// TIA Portal project "EMS" (V15.1) (continued)
   "Carrier_03_SitopSelectStatus" AT %I516.3 : Bool;   // SITOP SELECT STATUS
   "Carrier_03_DCsupplyOnPSCB2" AT %I516.4 : Bool;   // DC SUPPLY ON PSCB 2
   "Carrier_03_SpareInput(4_5)" AT %I516.5 : Bool;   // SPARE INPUT
   "Carrier_03_SpareInput(4_6)" AT %I516.6 : Bool;   // SPARE INPUT
   "Carrier_03_SpareInput(4_7)" AT %I516.7 : Bool;   // SPARE INPUT
   "Carrier_03_PB1_ProdHoldLH" AT %I517.0 : Bool;   // PB 1 PRODUCTION HOLD LH
   "Carrier_03_PB2_ResetLH" AT %I517.1 : Bool;   // PB 2 RESET LH
   "Carrier_03_PB3_ProdHoldRH" AT %I517.2 : Bool;   // PB 3 PRODUCTION HOLD RH
   "Carrier_03_PB4_ResetRH" AT %I517.3 : Bool;   // PB 4 RESET RH
   "Carrier_03_SpareInput(4_14)" AT %I517.4 : Bool;   // SPARE INPUT
   "Carrier_03_SpareInput(4_15)" AT %I517.5 : Bool;   // SPARE INPUT
   "Carrier_03_SpareInput(4_16)" AT %I517.6 : Bool;   // SPARE INPUT
   "Carrier_03_SpareInput(4_17)" AT %I517.7 : Bool;   // SPARE INPUT
   "Carrier_03_Slot5_Output" AT %IW518 : Word;   // SLOT 5 OUTPUT WORD
   "Carrier_03_IRD400_HMI_24VDC_ENABLE" AT %I518.0 : Bool;   // IRD 400 PANEL HMI 24V DC POWER
   "Carrier_03_FaultLight_LH" AT %I518.1 : Bool;   // FAULT LIGHT LH
   "Carrier_03_RunLight_LH" AT %I518.2 : Bool;   // RUN LIGHT LH
   "Carrier_03_FaultLight_RH" AT %I518.3 : Bool;   // FAULT LIGHT RH
   "Carrier_03_RunLight_RH" AT %I518.4 : Bool;   // RUN LIGHT RH
   "Carrier_03_SpareOutput(5_5)" AT %I518.5 : Bool;   // SPARE OUTPUT
   "Carrier_03_SpareOutput(5_6)" AT %I518.6 : Bool;   // SPARE OUTPUT
   "Carrier_03_SpareOutput(5_7)" AT %I518.7 : Bool;   // SPARE OUTPUT
   "Carrier_03_ActualSpeed" AT %IW520 : Word;   // ACTUAL SPEED
   "Carrier_03_CarrierDriveAlarm" AT %IW522 : Word;   // CARRIER DRIVE ALARM
   "Carrier_03_CarrierDriveWarning" AT %IW524 : Word;   // CARRIER DRIVE WARNING
   "Carrier_04_Status" AT %IW550 : Word;   // CARRIER STATUS WORD
   "Carrier_04_Status.0" AT %I550.0 : Bool;   // HEARTBEAT
   "Carrier_04_Status.1" AT %I550.1 : Bool;   // MANUAL
   "Carrier_04_Status.2" AT %I550.2 : Bool;   // IN_AUTO
   "Carrier_04_Status.3" AT %I550.3 : Bool;   // POSITIONING_COMPLETE
   "Carrier_04_Status.4" AT %I550.4 : Bool;   // PRODUCTION HOLD
   "Carrier_04_Status.5" AT %I550.5 : Bool;   // CARRIER MOVING FORWARD
   "Carrier_04_Status.6" AT %I550.6 : Bool;   // CARRIER MOVING REVERSE
   "Carrier_04_Status.7" AT %I550.7 : Bool;   // CARRIER FAULT
   "Carrier_04_Status.8" AT %I551.0 : Bool;   // CRASH DETECT TRIPPED
   "Carrier_04_Status.9" AT %I551.1 : Bool;
   "Carrier_04_Status.10" AT %I551.2 : Bool;
   "Carrier_04_Status.11" AT %I551.3 : Bool;
   "Carrier_04_Status.12" AT %I551.4 : Bool;
   "Carrier_04_Status.13" AT %I551.5 : Bool;
   "Carrier_04_Status.14" AT %I551.6 : Bool;
   "Carrier_04_Status.15" AT %I551.7 : Bool;
   "Carrier_04_SDCFaultCode" AT %IW552 : Word;   // SDC FAULT CODE
   "Carrier_04_CarrierPosition" AT %ID554 : DWord;   // CARRIER POSITION
   "Carrier_04_CarrierNumber" AT %IW558 : Word;   // CARRIER NUMBER
   "Carrier_04_G120DControlWord" AT %IW560 : Word;   // G120D_STW1_CONTROL
   "Carrier_04_G120DControlWord.0" AT %I560.0 : Bool;   // Bit_00_ON
   "Carrier_04_G120DControlWord.1" AT %I560.1 : Bool;   // Bit_01_AUS2_INH
   "Carrier_04_G120DControlWord.2" AT %I560.2 : Bool;   // Bit_02_AUS3_STOP
   "Carrier_04_G120DControlWord.3" AT %I560.3 : Bool;   // Bit_03_EN
   "Carrier_04_G120DControlWord.4" AT %I560.4 : Bool;   // Bit_04_EN_RAMP
   "Carrier_04_G120DControlWord.5" AT %I560.5 : Bool;   // Bit_05_START_RAMP
   "Carrier_04_G120DControlWord.6" AT %I560.6 : Bool;   // Bit_06_SETPOINT
   "Carrier_04_G120DControlWord.7" AT %I560.7 : Bool;   // Bit_07_RESET
   "Carrier_04_G120DControlWord.8" AT %I561.0 : Bool;   // Bit_08_JOG_R
   "Carrier_04_G120DControlWord.9" AT %I561.1 : Bool;   // Bit_09_JOG_L
   "Carrier_04_G120DControlWord.10" AT %I561.2 : Bool;   // Bit_10_CONTR_PLC
   "Carrier_04_G120DControlWord.11" AT %I561.3 : Bool;   // Bit_11_REVERSE
   "Carrier_04_G120DControlWord.12" AT %I561.4 : Bool;   // Bit_12_BRAKE_RELEASE
   "Carrier_04_G120DControlWord.13" AT %I561.5 : Bool;   // Bit_13_DDS
   "Carrier_04_G120DControlWord.14" AT %I561.6 : Bool;   // Bit_14_DO0
   "Carrier_04_G120DControlWord.15" AT %I561.7 : Bool;   // Bit_15_DO1
   "Carrier_04_G120DStatusWord" AT %IW562 : Word;   // G120D_ZSW1_STATUS
   "Carrier_04_G120DStatusWord.0" AT %I562.0 : Bool;   // Bit_00_READY_RUN
   "Carrier_04_G120DStatusWord.1" AT %I562.1 : Bool;   // Bit_01_READY_ON
   "Carrier_04_G120DStatusWord.2" AT %I562.2 : Bool;   // Bit_02_ENABLE
   "Carrier_04_G120DStatusWord.3" AT %I562.3 : Bool;   // Bit_03_FAULT
   "Carrier_04_G120DStatusWord.4" AT %I562.4 : Bool;   // Bit_04_OFF2
   "Carrier_04_G120DStatusWord.5" AT %I562.5 : Bool;   // Bit_05_OFF3
   "Carrier_04_G120DStatusWord.6" AT %I562.6 : Bool;   // Bit_06_LOCK_OUT
   "Carrier_04_G120DStatusWord.7" AT %I562.7 : Bool;   // Bit_07_WARN
   "Carrier_04_G120DStatusWord.8" AT %I563.0 : Bool;   // Bit_08_NO_DEVIATION
   "Carrier_04_G120DStatusWord.9" AT %I563.1 : Bool;   // Bit_09_CONTR_PLC
   "Carrier_04_G120DStatusWord.10" AT %I563.2 : Bool;   // Bit_10_F_MAX
   "Carrier_04_G120DStatusWord.11" AT %I563.3 : Bool;   // Bit_11_LIMIT_REACHED
   "Carrier_04_G120DStatusWord.12" AT %I563.4 : Bool;   // Bit_12_BRAKE_OPEN
   "Carrier_04_G120DStatusWord.13" AT %I563.5 : Bool;   // Bit_13_NO_OVERTEMP
   "Carrier_04_G120DStatusWord.14" AT %I563.6 : Bool;   // Bit_14_CW_CCW
   "Carrier_04_G120DStatusWord.15" AT %I563.7 : Bool;   // Bit_15_OVERL
   "Carrier_04_Slot2_Input" AT %IW564 : Word;   // SLOT 2 INPUT WORD
   "Carrier_04_CrashDetectSW" AT %I564.0 : Bool;   // CRASH DETECT SW
   "Carrier_04_SpareSafetyInput(2_1)" AT %I564.1 : Bool;   // SPARE SAFETY INPUT
   "Carrier_04_SpareSafetyInput(2_2)" AT %I564.2 : Bool;   // SPARE SAFETY INPUT
   "Carrier_04_SpareSafetyInput(2_3)" AT %I564.3 : Bool;   // SPARE SAFETY INPUT
   "Carrier_04_SpareSafetyInput(2_4)" AT %I564.4 : Bool;   // SPARE SAFETY INPUT
   "Carrier_04_SpareSafetyInput(2_5)" AT %I564.5 : Bool;   // SPARE SAFETY INPUT
   "Carrier_04_SpareSafetyInput(2_6)" AT %I564.6 : Bool;   // SPARE SAFETY INPUT
   "Carrier_04_SpareSafetyInput(2_7)" AT %I564.7 : Bool;   // SPARE SAFETY INPUT
   "Carrier_04_Slot3_SafetyOutput" AT %IW565 : Word;   // SLOT 3 SAFETY OUTPUT WORD
   "Carrier_04_Crash_Detect_OK" AT %I565.0 : Bool;   // CARRIER CRASH DETECT
   "Carrier_04_SpareSafetyOutput(3_1)" AT %I565.1 : Bool;   // SPARE SAFETY OUTPUT
   "Carrier_04_SpareSafetyOutput(3_2)" AT %I565.2 : Bool;   // SPARE SAFETY OUTPUT
   "Carrier_04_SpareSafetyOutput(3_3)" AT %I565.3 : Bool;   // SPARE SAFETY OUTPUT
   "Carrier_04_SpareSafetyOutput(3_4)" AT %I565.4 : Bool;   // SPARE SAFETY OUTPUT
   "Carrier_04_SpareSafetyOutput(3_5)" AT %I565.5 : Bool;   // SPARE SAFETY OUTPUT
   "Carrier_04_SpareSafetyOutput(3_6)" AT %I565.6 : Bool;   // SPARE SAFETY OUTPUT
   "Carrier_04_SpareSafetyOutput(3_7)" AT %I565.7 : Bool;   // SPARE SAFETY OUTPUT
   "Carrier_04_Slot4_Input" AT %IW566 : Word;   // SLOT 4 INPUT WORD
   "Carrier_04_480VPowerOn_MDCB1" AT %I566.0 : Bool;   // 480 VAC POWER ON MDCB 1
   "Carrier_04_SpareInput(4_1)" AT %I566.1 : Bool;   // SPARE INPUT
   "Carrier_04_SpareInput(4_2)" AT %I566.2 : Bool;   // SPARE INPUT
   "Carrier_04_SitopSelectStatus" AT %I566.3 : Bool;   // SITOP SELECT STATUS
   "Carrier_04_DCsupplyOnPSCB2" AT %I566.4 : Bool;   // DC SUPPLY ON PSCB 2
   "Carrier_04_SpareInput(4_5)" AT %I566.5 : Bool;   // SPARE INPUT
   "Carrier_04_SpareInput(4_6)" AT %I566.6 : Bool;   // SPARE INPUT
   "Carrier_04_SpareInput(4_7)" AT %I566.7 : Bool;   // SPARE INPUT
   "Carrier_04_PB1_ProdHoldLH" AT %I567.0 : Bool;   // PB 1 PRODUCTION HOLD LH
   "Carrier_04_PB2_ResetLH" AT %I567.1 : Bool;   // PB 2 RESET LH
   "Carrier_04_PB3_ProdHoldRH" AT %I567.2 : Bool;   // PB 3 PRODUCTION HOLD RH
   "Carrier_04_PB4_ResetRH" AT %I567.3 : Bool;   // PB 4 RESET RH
   "Carrier_04_SpareInput(4_14)" AT %I567.4 : Bool;   // SPARE INPUT
   "Carrier_04_SpareInput(4_15)" AT %I567.5 : Bool;   // SPARE INPUT
   "Carrier_04_SpareInput(4_16)" AT %I567.6 : Bool;   // SPARE INPUT
   "Carrier_04_SpareInput(4_17)" AT %I567.7 : Bool;   // SPARE INPUT
   "Carrier_04_Slot5_Output" AT %IW568 : Word;   // SLOT 5 OUTPUT WORD
   "Carrier_04_IRD400_HMI_24VDC_ENABLE" AT %I568.0 : Bool;   // IRD 400 PANEL HMI 24V DC POWER
   "Carrier_04_FaultLight_LH" AT %I568.1 : Bool;   // FAULT LIGHT LH
   "Carrier_04_RunLight_LH" AT %I568.2 : Bool;   // RUN LIGHT LH
   "Carrier_04_FaultLight_RH" AT %I568.3 : Bool;   // FAULT LIGHT RH
   "Carrier_04_RunLight_RH" AT %I568.4 : Bool;   // RUN LIGHT RH
   "Carrier_04_SpareOutput(5_5)" AT %I568.5 : Bool;   // SPARE OUTPUT
   "Carrier_04_SpareOutput(5_6)" AT %I568.6 : Bool;   // SPARE OUTPUT
   "Carrier_04_SpareOutput(5_7)" AT %I568.7 : Bool;   // SPARE OUTPUT
   "Carrier_04_ActualSpeed" AT %IW570 : Word;   // ACTUAL SPEED
   "Carrier_04_CarrierDriveAlarm" AT %IW572 : Word;   // CARRIER DRIVE ALARM
   "Carrier_04_CarrierDriveWarning" AT %IW574 : Word;   // CARRIER DRIVE WARNING
   "Carrier_05_Status" AT %IW600 : Word;   // CARRIER STATUS WORD
   "Carrier_05_Status.0" AT %I600.0 : Bool;   // HEARTBEAT
   "Carrier_05_Status.1" AT %I600.1 : Bool;   // MANUAL
   "Carrier_05_Status.2" AT %I600.2 : Bool;   // IN_AUTO
   "Carrier_05_Status.3" AT %I600.3 : Bool;   // POSITIONING_COMPLETE
   "Carrier_05_Status.4" AT %I600.4 : Bool;   // PRODUCTION HOLD
   "Carrier_05_Status.5" AT %I600.5 : Bool;   // CARRIER MOVING FORWARD
   "Carrier_05_Status.6" AT %I600.6 : Bool;   // CARRIER MOVING REVERSE
   "Carrier_05_Status.7" AT %I600.7 : Bool;   // CARRIER FAULT
   "Carrier_05_Status.8" AT %I601.0 : Bool;   // CRASH DETECT TRIPPED
   "Carrier_05_Status.9" AT %I601.1 : Bool;
   "Carrier_05_Status.10" AT %I601.2 : Bool;
   "Carrier_05_Status.11" AT %I601.3 : Bool;
   "Carrier_05_Status.12" AT %I601.4 : Bool;
   "Carrier_05_Status.13" AT %I601.5 : Bool;
   "Carrier_05_Status.14" AT %I601.6 : Bool;
   "Carrier_05_Status.15" AT %I601.7 : Bool;
   "Carrier_05_SDCFaultCode" AT %IW602 : Word;   // SDC FAULT CODE
   "Carrier_05_CarrierPosition" AT %ID604 : DWord;   // CARRIER POSITION
   "Carrier_05_CarrierNumber" AT %IW608 : Word;   // CARRIER NUMBER
   "Carrier_05_G120DControlWord" AT %IW610 : Word;   // G120D_STW1_CONTROL
   "Carrier_05_G120DControlWord.0" AT %I610.0 : Bool;   // Bit_00_ON
   "Carrier_05_G120DControlWord.1" AT %I610.1 : Bool;   // Bit_01_AUS2_INH
   "Carrier_05_G120DControlWord.2" AT %I610.2 : Bool;   // Bit_02_AUS3_STOP
   "Carrier_05_G120DControlWord.3" AT %I610.3 : Bool;   // Bit_03_EN
   "Carrier_05_G120DControlWord.4" AT %I610.4 : Bool;   // Bit_04_EN_RAMP
   "Carrier_05_G120DControlWord.5" AT %I610.5 : Bool;   // Bit_05_START_RAMP
   "Carrier_05_G120DControlWord.6" AT %I610.6 : Bool;   // Bit_06_SETPOINT
   "Carrier_05_G120DControlWord.7" AT %I610.7 : Bool;   // Bit_07_RESET
   "Carrier_05_G120DControlWord.8" AT %I611.0 : Bool;   // Bit_08_JOG_R
   "Carrier_05_G120DControlWord.9" AT %I611.1 : Bool;   // Bit_09_JOG_L
   "Carrier_05_G120DControlWord.10" AT %I611.2 : Bool;   // Bit_10_CONTR_PLC
   "Carrier_05_G120DControlWord.11" AT %I611.3 : Bool;   // Bit_11_REVERSE
   "Carrier_05_G120DControlWord.12" AT %I611.4 : Bool;   // Bit_12_BRAKE_RELEASE
   "Carrier_05_G120DControlWord.13" AT %I611.5 : Bool;   // Bit_13_DDS
   "Carrier_05_G120DControlWord.14" AT %I611.6 : Bool;   // Bit_14_DO0
   "Carrier_05_G120DControlWord.15" AT %I611.7 : Bool;   // Bit_15_DO1
   "Carrier_05_G120DStatusWord" AT %IW612 : Word;   // G120D_ZSW1_STATUS
   "Carrier_05_G120DStatusWord.0" AT %I612.0 : Bool;   // Bit_00_READY_RUN
   "Carrier_05_G120DStatusWord.1" AT %I612.1 : Bool;   // Bit_01_READY_ON
   "Carrier_05_G120DStatusWord.2" AT %I612.2 : Bool;   // Bit_02_ENABLE
   "Carrier_05_G120DStatusWord.3" AT %I612.3 : Bool;   // Bit_03_FAULT
   "Carrier_05_G120DStatusWord.4" AT %I612.4 : Bool;   // Bit_04_OFF2
   "Carrier_05_G120DStatusWord.5" AT %I612.5 : Bool;   // Bit_05_OFF3
   "Carrier_05_G120DStatusWord.6" AT %I612.6 : Bool;   // Bit_06_LOCK_OUT
   "Carrier_05_G120DStatusWord.7" AT %I612.7 : Bool;   // Bit_07_WARN
   "Carrier_05_G120DStatusWord.8" AT %I613.0 : Bool;   // Bit_08_NO_DEVIATION
   "Carrier_05_G120DStatusWord.9" AT %I613.1 : Bool;   // Bit_09_CONTR_PLC
   "Carrier_05_G120DStatusWord.10" AT %I613.2 : Bool;   // Bit_10_F_MAX
   "Carrier_05_G120DStatusWord.11" AT %I613.3 : Bool;   // Bit_11_LIMIT_REACHED
   "Carrier_05_G120DStatusWord.12" AT %I613.4 : Bool;   // Bit_12_BRAKE_OPEN
   "Carrier_05_G120DStatusWord.13" AT %I613.5 : Bool;   // Bit_13_NO_OVERTEMP
   "Carrier_05_G120DStatusWord.14" AT %I613.6 : Bool;   // Bit_14_CW_CCW
   "Carrier_05_G120DStatusWord.15" AT %I613.7 : Bool;   // Bit_15_OVERL
   "Carrier_05_Slot2_Input" AT %IW614 : Word;   // SLOT 2 INPUT WORD
   "Carrier_05_CrashDetectSW" AT %I614.0 : Bool;   // CRASH DETECT SW
   "Carrier_05_SpareSafetyInput(2_1)" AT %I614.1 : Bool;   // SPARE SAFETY INPUT
   "Carrier_05_SpareSafetyInput(2_2)" AT %I614.2 : Bool;   // SPARE SAFETY INPUT
   "Carrier_05_SpareSafetyInput(2_3)" AT %I614.3 : Bool;   // SPARE SAFETY INPUT
   "Carrier_05_SpareSafetyInput(2_4)" AT %I614.4 : Bool;   // SPARE SAFETY INPUT
   "Carrier_05_SpareSafetyInput(2_5)" AT %I614.5 : Bool;   // SPARE SAFETY INPUT
   "Carrier_05_SpareSafetyInput(2_6)" AT %I614.6 : Bool;   // SPARE SAFETY INPUT
   "Carrier_05_SpareSafetyInput(2_7)" AT %I614.7 : Bool;   // SPARE SAFETY INPUT
   "Carrier_05_Slot3_SafetyOutput" AT %IW615 : Word;   // SLOT 3 SAFETY OUTPUT WORD
   "Carrier_05_Crash_Detect_OK" AT %I615.0 : Bool;   // CARRIER CRASH DETECT
   "Carrier_05_SpareSafetyOutput(3_1)" AT %I615.1 : Bool;   // SPARE SAFETY OUTPUT
   "Carrier_05_SpareSafetyOutput(3_2)" AT %I615.2 : Bool;   // SPARE SAFETY OUTPUT
   "Carrier_05_SpareSafetyOutput(3_3)" AT %I615.3 : Bool;   // SPARE SAFETY OUTPUT
   "Carrier_05_SpareSafetyOutput(3_4)" AT %I615.4 : Bool;   // SPARE SAFETY OUTPUT
   "Carrier_05_SpareSafetyOutput(3_5)" AT %I615.5 : Bool;   // SPARE SAFETY OUTPUT
   "Carrier_05_SpareSafetyOutput(3_6)" AT %I615.6 : Bool;   // SPARE SAFETY OUTPUT
   "Carrier_05_SpareSafetyOutput(3_7)" AT %I615.7 : Bool;   // SPARE SAFETY OUTPUT
   "Carrier_05_Slot4_Input" AT %IW616 : Word;   // SLOT 4 INPUT WORD
   "Carrier_05_480VPowerOn_MDCB1" AT %I616.0 : Bool;   // 480 VAC POWER ON MDCB 1
   "Carrier_05_SpareInput(4_1)" AT %I616.1 : Bool;   // SPARE INPUT
   "Carrier_05_SpareInput(4_2)" AT %I616.2 : Bool;   // SPARE INPUT
   "Carrier_05_SitopSelectStatus" AT %I616.3 : Bool;   // SITOP SELECT STATUS
   "Carrier_05_DCsupplyOnPSCB2" AT %I616.4 : Bool;   // DC SUPPLY ON PSCB 2
   "Carrier_05_SpareInput(4_5)" AT %I616.5 : Bool;   // SPARE INPUT
   "Carrier_05_SpareInput(4_6)" AT %I616.6 : Bool;   // SPARE INPUT
   "Carrier_05_SpareInput(4_7)" AT %I616.7 : Bool;   // SPARE INPUT
   "Carrier_05_PB1_ProdHoldLH" AT %I617.0 : Bool;   // PB 1 PRODUCTION HOLD LH
   "Carrier_05_PB2_ResetLH" AT %I617.1 : Bool;   // PB 2 RESET LH
   "Carrier_05_PB3_ProdHoldRH" AT %I617.2 : Bool;   // PB 3 PRODUCTION HOLD RH
   "Carrier_05_PB4_ResetRH" AT %I617.3 : Bool;   // PB 4 RESET RH
   "Carrier_05_SpareInput(4_14)" AT %I617.4 : Bool;   // SPARE INPUT
   "Carrier_05_SpareInput(4_15)" AT %I617.5 : Bool;   // SPARE INPUT
   "Carrier_05_SpareInput(4_16)" AT %I617.6 : Bool;   // SPARE INPUT
   "Carrier_05_SpareInput(4_17)" AT %I617.7 : Bool;   // SPARE INPUT
   "Carrier_05_Slot5_Output" AT %IW618 : Word;   // SLOT 5 OUTPUT WORD
   "Carrier_05_IRD400_HMI_24VDC_ENABLE" AT %I618.0 : Bool;   // IRD 400 PANEL HMI 24V DC POWER
   "Carrier_05_FaultLight_LH" AT %I618.1 : Bool;   // FAULT LIGHT LH
   "Carrier_05_RunLight_LH" AT %I618.2 : Bool;   // RUN LIGHT LH
   "Carrier_05_FaultLight_RH" AT %I618.3 : Bool;   // FAULT LIGHT RH
   "Carrier_05_RunLight_RH" AT %I618.4 : Bool;   // RUN LIGHT RH
   "Carrier_05_SpareOutput(5_5)" AT %I618.5 : Bool;   // SPARE OUTPUT
   "Carrier_05_SpareOutput(5_6)" AT %I618.6 : Bool;   // SPARE OUTPUT
   "Carrier_05_SpareOutput(5_7)" AT %I618.7 : Bool;   // SPARE OUTPUT
   "Carrier_05_ActualSpeed" AT %IW620 : Word;   // ACTUAL SPEED
   "Carrier_05_CarrierDriveAlarm" AT %IW622 : Word;   // CARRIER DRIVE ALARM
   "Carrier_05_CarrierDriveWarning" AT %IW624 : Word;   // CARRIER DRIVE WARNING
   "Carrier_06_Status" AT %IW650 : Word;   // CARRIER STATUS WORD
   "Carrier_06_Status.0" AT %I650.0 : Bool;   // HEARTBEAT
   "Carrier_06_Status.1" AT %I650.1 : Bool;   // MANUAL
   "Carrier_06_Status.2" AT %I650.2 : Bool;   // IN_AUTO
   "Carrier_06_Status.3" AT %I650.3 : Bool;   // POSITIONING_COMPLETE
   "Carrier_06_Status.4" AT %I650.4 : Bool;   // PRODUCTION HOLD
   "Carrier_06_Status.5" AT %I650.5 : Bool;   // CARRIER MOVING FORWARD
   "Carrier_06_Status.6" AT %I650.6 : Bool;   // CARRIER MOVING REVERSE
   "Carrier_06_Status.7" AT %I650.7 : Bool;   // CARRIER FAULT
   "Carrier_06_Status.8" AT %I651.0 : Bool;   // CRASH DETECT TRIPPED
   "Carrier_06_Status.9" AT %I651.1 : Bool;
   "Carrier_06_Status.10" AT %I651.2 : Bool;
   "Carrier_06_Status.11" AT %I651.3 : Bool;
   "Carrier_06_Status.12" AT %I651.4 : Bool;
   "Carrier_06_Status.13" AT %I651.5 : Bool;
   "Carrier_06_Status.14" AT %I651.6 : Bool;
   "Carrier_06_Status.15" AT %I651.7 : Bool;
   "Carrier_06_SDCFaultCode" AT %IW652 : Word;   // SDC FAULT CODE
   "Carrier_06_CarrierPosition" AT %ID654 : DWord;   // CARRIER POSITION
   "Carrier_06_CarrierNumber" AT %IW658 : Word;   // CARRIER NUMBER
   "Carrier_06_G120DControlWord" AT %IW660 : Word;   // G120D_STW1_CONTROL
   "Carrier_06_G120DControlWord.0" AT %I660.0 : Bool;   // Bit_00_ON
   "Carrier_06_G120DControlWord.1" AT %I660.1 : Bool;   // Bit_01_AUS2_INH
   "Carrier_06_G120DControlWord.2" AT %I660.2 : Bool;   // Bit_02_AUS3_STOP
   "Carrier_06_G120DControlWord.3" AT %I660.3 : Bool;   // Bit_03_EN
   "Carrier_06_G120DControlWord.4" AT %I660.4 : Bool;   // Bit_04_EN_RAMP
   "Carrier_06_G120DControlWord.5" AT %I660.5 : Bool;   // Bit_05_START_RAMP
   "Carrier_06_G120DControlWord.6" AT %I660.6 : Bool;   // Bit_06_SETPOINT
   "Carrier_06_G120DControlWord.7" AT %I660.7 : Bool;   // Bit_07_RESET
   "Carrier_06_G120DControlWord.8" AT %I661.0 : Bool;   // Bit_08_JOG_R
   "Carrier_06_G120DControlWord.9" AT %I661.1 : Bool;   // Bit_09_JOG_L
   "Carrier_06_G120DControlWord.10" AT %I661.2 : Bool;   // Bit_10_CONTR_PLC
   "Carrier_06_G120DControlWord.11" AT %I661.3 : Bool;   // Bit_11_REVERSE
   "Carrier_06_G120DControlWord.12" AT %I661.4 : Bool;   // Bit_12_BRAKE_RELEASE
   "Carrier_06_G120DControlWord.13" AT %I661.5 : Bool;   // Bit_13_DDS
   "Carrier_06_G120DControlWord.14" AT %I661.6 : Bool;   // Bit_14_DO0
   "Carrier_06_G120DControlWord.15" AT %I661.7 : Bool;   // Bit_15_DO1
   "Carrier_06_G120DStatusWord" AT %IW662 : Word;   // G120D_ZSW1_STATUS
   "Carrier_06_G120DStatusWord.0" AT %I662.0 : Bool;   // Bit_00_READY_RUN
   "Carrier_06_G120DStatusWord.1" AT %I662.1 : Bool;   // Bit_01_READY_ON
   "Carrier_06_G120DStatusWord.2" AT %I662.2 : Bool;   // Bit_02_ENABLE
   "Carrier_06_G120DStatusWord.3" AT %I662.3 : Bool;   // Bit_03_FAULT
   "Carrier_06_G120DStatusWord.4" AT %I662.4 : Bool;   // Bit_04_OFF2
   "Carrier_06_G120DStatusWord.5" AT %I662.5 : Bool;   // Bit_05_OFF3
   "Carrier_06_G120DStatusWord.6" AT %I662.6 : Bool;   // Bit_06_LOCK_OUT
   "Carrier_06_G120DStatusWord.7" AT %I662.7 : Bool;   // Bit_07_WARN
   "Carrier_06_G120DStatusWord.8" AT %I663.0 : Bool;   // Bit_08_NO_DEVIATION
   "Carrier_06_G120DStatusWord.9" AT %I663.1 : Bool;   // Bit_09_CONTR_PLC
   "Carrier_06_G120DStatusWord.10" AT %I663.2 : Bool;   // Bit_10_F_MAX
   "Carrier_06_G120DStatusWord.11" AT %I663.3 : Bool;   // Bit_11_LIMIT_REACHED
   "Carrier_06_G120DStatusWord.12" AT %I663.4 : Bool;   // Bit_12_BRAKE_OPEN
   "Carrier_06_G120DStatusWord.13" AT %I663.5 : Bool;   // Bit_13_NO_OVERTEMP
   "Carrier_06_G120DStatusWord.14" AT %I663.6 : Bool;   // Bit_14_CW_CCW
   "Carrier_06_G120DStatusWord.15" AT %I663.7 : Bool;   // Bit_15_OVERL
   "Carrier_06_Slot2_Input" AT %IW664 : Word;   // SLOT 2 INPUT WORD
   "Carrier_06_CrashDetectSW" AT %I664.0 : Bool;   // CRASH DETECT SW
   "Carrier_06_SpareSafetyInput(2_1)" AT %I664.1 : Bool;   // SPARE SAFETY INPUT
   "Carrier_06_SpareSafetyInput(2_2)" AT %I664.2 : Bool;   // SPARE SAFETY INPUT
   "Carrier_06_SpareSafetyInput(2_3)" AT %I664.3 : Bool;   // SPARE SAFETY INPUT
   "Carrier_06_SpareSafetyInput(2_4)" AT %I664.4 : Bool;   // SPARE SAFETY INPUT
   "Carrier_06_SpareSafetyInput(2_5)" AT %I664.5 : Bool;   // SPARE SAFETY INPUT
   "Carrier_06_SpareSafetyInput(2_6)" AT %I664.6 : Bool;   // SPARE SAFETY INPUT
   "Carrier_06_SpareSafetyInput(2_7)" AT %I664.7 : Bool;   // SPARE SAFETY INPUT
   "Carrier_06_Slot3_SafetyOutput" AT %IW665 : Word;   // SLOT 3 SAFETY OUTPUT WORD
   "Carrier_06_Crash_Detect_OK" AT %I665.0 : Bool;   // CARRIER CRASH DETECT
   "Carrier_06_SpareSafetyOutput(3_1)" AT %I665.1 : Bool;   // SPARE SAFETY OUTPUT
   "Carrier_06_SpareSafetyOutput(3_2)" AT %I665.2 : Bool;   // SPARE SAFETY OUTPUT
   "Carrier_06_SpareSafetyOutput(3_3)" AT %I665.3 : Bool;   // SPARE SAFETY OUTPUT
   "Carrier_06_SpareSafetyOutput(3_4)" AT %I665.4 : Bool;   // SPARE SAFETY OUTPUT
   "Carrier_06_SpareSafetyOutput(3_5)" AT %I665.5 : Bool;   // SPARE SAFETY OUTPUT
   "Carrier_06_SpareSafetyOutput(3_6)" AT %I665.6 : Bool;   // SPARE SAFETY OUTPUT
   "Carrier_06_SpareSafetyOutput(3_7)" AT %I665.7 : Bool;   // SPARE SAFETY OUTPUT
   "Carrier_06_Slot4_Input" AT %IW666 : Word;   // SLOT 4 INPUT WORD
   "Carrier_06_480VPowerOn_MDCB1" AT %I666.0 : Bool;   // 480 VAC POWER ON MDCB 1
   "Carrier_06_SpareInput(4_1)" AT %I666.1 : Bool;   // SPARE INPUT
   "Carrier_06_SpareInput(4_2)" AT %I666.2 : Bool;   // SPARE INPUT
   "Carrier_06_SitopSelectStatus" AT %I666.3 : Bool;   // SITOP SELECT STATUS
   "Carrier_06_DCsupplyOnPSCB2" AT %I666.4 : Bool;   // DC SUPPLY ON PSCB 2
   "Carrier_06_SpareInput(4_5)" AT %I666.5 : Bool;   // SPARE INPUT
   "Carrier_06_SpareInput(4_6)" AT %I666.6 : Bool;   // SPARE INPUT
   "Carrier_06_SpareInput(4_7)" AT %I666.7 : Bool;   // SPARE INPUT
   "Carrier_06_PB1_ProdHoldLH" AT %I667.0 : Bool;   // PB 1 PRODUCTION HOLD LH
   "Carrier_06_PB2_ResetLH" AT %I667.1 : Bool;   // PB 2 RESET LH
   "Carrier_06_PB3_ProdHoldRH" AT %I667.2 : Bool;   // PB 3 PRODUCTION HOLD RH
   "Carrier_06_PB4_ResetRH" AT %I667.3 : Bool;   // PB 4 RESET RH
   "Carrier_06_SpareInput(4_14)" AT %I667.4 : Bool;   // SPARE INPUT
   "Carrier_06_SpareInput(4_15)" AT %I667.5 : Bool;   // SPARE INPUT
   "Carrier_06_SpareInput(4_16)" AT %I667.6 : Bool;   // SPARE INPUT
   "Carrier_06_SpareInput(4_17)" AT %I667.7 : Bool;   // SPARE INPUT
   "Carrier_06_Slot5_Output" AT %IW668 : Word;   // SLOT 5 OUTPUT WORD
   "Carrier_06_IRD400_HMI_24VDC_ENABLE" AT %I668.0 : Bool;   // IRD 400 PANEL HMI 24V DC POWER
   "Carrier_06_FaultLight_LH" AT %I668.1 : Bool;   // FAULT LIGHT LH
   "Carrier_06_RunLight_LH" AT %I668.2 : Bool;   // RUN LIGHT LH
   "Carrier_06_FaultLight_RH" AT %I668.3 : Bool;   // FAULT LIGHT RH
   "Carrier_06_RunLight_RH" AT %I668.4 : Bool;   // RUN LIGHT RH
   "Carrier_06_SpareOutput(5_5)" AT %I668.5 : Bool;   // SPARE OUTPUT
   "Carrier_06_SpareOutput(5_6)" AT %I668.6 : Bool;   // SPARE OUTPUT
   "Carrier_06_SpareOutput(5_7)" AT %I668.7 : Bool;   // SPARE OUTPUT
   "Carrier_06_ActualSpeed" AT %IW670 : Word;   // ACTUAL SPEED
   "Carrier_06_CarrierDriveAlarm" AT %IW672 : Word;   // CARRIER DRIVE ALARM
   "Carrier_06_CarrierDriveWarning" AT %IW674 : Word;   // CARRIER DRIVE WARNING
   "Carrier_07_Status" AT %IW700 : Word;   // CARRIER STATUS WORD
   "Carrier_07_Status.0" AT %I700.0 : Bool;   // HEARTBEAT
   "Carrier_07_Status.1" AT %I700.1 : Bool;   // MANUAL
   "Carrier_07_Status.2" AT %I700.2 : Bool;   // IN_AUTO
   "Carrier_07_Status.3" AT %I700.3 : Bool;   // POSITIONING_COMPLETE
   "Carrier_07_Status.4" AT %I700.4 : Bool;   // PRODUCTION HOLD
   "Carrier_07_Status.5" AT %I700.5 : Bool;   // CARRIER MOVING FORWARD
   "Carrier_07_Status.6" AT %I700.6 : Bool;   // CARRIER MOVING REVERSE
   "Carrier_07_Status.7" AT %I700.7 : Bool;   // CARRIER FAULT
   "Carrier_07_Status.8" AT %I701.0 : Bool;   // CRASH DETECT TRIPPED
   "Carrier_07_Status.9" AT %I701.1 : Bool;
   "Carrier_07_Status.10" AT %I701.2 : Bool;
   "Carrier_07_Status.11" AT %I701.3 : Bool;
   "Carrier_07_Status.12" AT %I701.4 : Bool;
   "Carrier_07_Status.13" AT %I701.5 : Bool;
   "Carrier_07_Status.14" AT %I701.6 : Bool;
   "Carrier_07_Status.15" AT %I701.7 : Bool;
   "Carrier_07_SDCFaultCode" AT %IW702 : Word;   // SDC FAULT CODE
   "Carrier_07_CarrierPosition" AT %ID704 : DWord;   // CARRIER POSITION
   "Carrier_07_CarrierNumber" AT %IW708 : Word;   // CARRIER NUMBER
   "Carrier_07_G120DControlWord" AT %IW710 : Word;   // G120D_STW1_CONTROL
   "Carrier_07_G120DControlWord.0" AT %I710.0 : Bool;   // Bit_00_ON
   "Carrier_07_G120DControlWord.1" AT %I710.1 : Bool;   // Bit_01_AUS2_INH
   "Carrier_07_G120DControlWord.2" AT %I710.2 : Bool;   // Bit_02_AUS3_STOP
   "Carrier_07_G120DControlWord.3" AT %I710.3 : Bool;   // Bit_03_EN
   "Carrier_07_G120DControlWord.4" AT %I710.4 : Bool;   // Bit_04_EN_RAMP
   "Carrier_07_G120DControlWord.5" AT %I710.5 : Bool;   // Bit_05_START_RAMP
   "Carrier_07_G120DControlWord.6" AT %I710.6 : Bool;   // Bit_06_SETPOINT
   "Carrier_07_G120DControlWord.7" AT %I710.7 : Bool;   // Bit_07_RESET
   "Carrier_07_G120DControlWord.8" AT %I711.0 : Bool;   // Bit_08_JOG_R
   "Carrier_07_G120DControlWord.9" AT %I711.1 : Bool;   // Bit_09_JOG_L
   "Carrier_07_G120DControlWord.10" AT %I711.2 : Bool;   // Bit_10_CONTR_PLC
   "Carrier_07_G120DControlWord.11" AT %I711.3 : Bool;   // Bit_11_REVERSE
   "Carrier_07_G120DControlWord.12" AT %I711.4 : Bool;   // Bit_12_BRAKE_RELEASE
   "Carrier_07_G120DControlWord.13" AT %I711.5 : Bool;   // Bit_13_DDS
   "Carrier_07_G120DControlWord.14" AT %I711.6 : Bool;   // Bit_14_DO0
   "Carrier_07_G120DControlWord.15" AT %I711.7 : Bool;   // Bit_15_DO1
   "Carrier_07_G120DStatusWord" AT %IW712 : Word;   // G120D_ZSW1_STATUS
   "Carrier_07_G120DStatusWord.0" AT %I712.0 : Bool;   // Bit_00_READY_RUN
   "Carrier_07_G120DStatusWord.1" AT %I712.1 : Bool;   // Bit_01_READY_ON
   "Carrier_07_G120DStatusWord.2" AT %I712.2 : Bool;   // Bit_02_ENABLE
   "Carrier_07_G120DStatusWord.3" AT %I712.3 : Bool;   // Bit_03_FAULT
   "Carrier_07_G120DStatusWord.4" AT %I712.4 : Bool;   // Bit_04_OFF2
   "Carrier_07_G120DStatusWord.5" AT %I712.5 : Bool;   // Bit_05_OFF3
   "Carrier_07_G120DStatusWord.6" AT %I712.6 : Bool;   // Bit_06_LOCK_OUT
   "Carrier_07_G120DStatusWord.7" AT %I712.7 : Bool;   // Bit_07_WARN
   "Carrier_07_G120DStatusWord.8" AT %I713.0 : Bool;   // Bit_08_NO_DEVIATION
   "Carrier_07_G120DStatusWord.9" AT %I713.1 : Bool;   // Bit_09_CONTR_PLC
   "Carrier_07_G120DStatusWord.10" AT %I713.2 : Bool;   // Bit_10_F_MAX
   "Carrier_07_G120DStatusWord.11" AT %I713.3 : Bool;   // Bit_11_LIMIT_REACHED
   "Carrier_07_G120DStatusWord.12" AT %I713.4 : Bool;   // Bit_12_BRAKE_OPEN
   "Carrier_07_G120DStatusWord.13" AT %I713.5 : Bool;   // Bit_13_NO_OVERTEMP
   "Carrier_07_G120DStatusWord.14" AT %I713.6 : Bool;   // Bit_14_CW_CCW
   "Carrier_07_G120DStatusWord.15" AT %I713.7 : Bool;   // Bit_15_OVERL
   "Carrier_07_Slot2_Input" AT %IW714 : Word;   // SLOT 2 INPUT WORD
   "Carrier_07_CrashDetectSW" AT %I714.0 : Bool;   // CRASH DETECT SW
   "Carrier_07_SpareSafetyInput(2_1)" AT %I714.1 : Bool;   // SPARE SAFETY INPUT
   "Carrier_07_SpareSafetyInput(2_2)" AT %I714.2 : Bool;   // SPARE SAFETY INPUT
   "Carrier_07_SpareSafetyInput(2_3)" AT %I714.3 : Bool;   // SPARE SAFETY INPUT
   "Carrier_07_SpareSafetyInput(2_4)" AT %I714.4 : Bool;   // SPARE SAFETY INPUT
   "Carrier_07_SpareSafetyInput(2_5)" AT %I714.5 : Bool;   // SPARE SAFETY INPUT
   "Carrier_07_SpareSafetyInput(2_6)" AT %I714.6 : Bool;   // SPARE SAFETY INPUT
   "Carrier_07_SpareSafetyInput(2_7)" AT %I714.7 : Bool;   // SPARE SAFETY INPUT
   "Carrier_07_Slot3_SafetyOutput" AT %IW715 : Word;   // SLOT 3 SAFETY OUTPUT WORD
   "Carrier_07_Crash_Detect_OK" AT %I715.0 : Bool;   // CARRIER CRASH DETECT
   "Carrier_07_SpareSafetyOutput(3_1)" AT %I715.1 : Bool;   // SPARE SAFETY OUTPUT
   "Carrier_07_SpareSafetyOutput(3_2)" AT %I715.2 : Bool;   // SPARE SAFETY OUTPUT
   "Carrier_07_SpareSafetyOutput(3_3)" AT %I715.3 : Bool;   // SPARE SAFETY OUTPUT
   "Carrier_07_SpareSafetyOutput(3_4)" AT %I715.4 : Bool;   // SPARE SAFETY OUTPUT
   "Carrier_07_SpareSafetyOutput(3_5)" AT %I715.5 : Bool;   // SPARE SAFETY OUTPUT
   "Carrier_07_SpareSafetyOutput(3_6)" AT %I715.6 : Bool;   // SPARE SAFETY OUTPUT
   "Carrier_07_SpareSafetyOutput(3_7)" AT %I715.7 : Bool;   // SPARE SAFETY OUTPUT
   "Carrier_07_Slot4_Input" AT %IW716 : Word;   // SLOT 4 INPUT WORD
   "Carrier_07_480VPowerOn_MDCB1" AT %I716.0 : Bool;   // 480 VAC POWER ON MDCB 1
   "Carrier_07_SpareInput(4_1)" AT %I716.1 : Bool;   // SPARE INPUT
   "Carrier_07_SpareInput(4_2)" AT %I716.2 : Bool;   // SPARE INPUT
   "Carrier_07_SitopSelectStatus" AT %I716.3 : Bool;   // SITOP SELECT STATUS
   "Carrier_07_DCsupplyOnPSCB2" AT %I716.4 : Bool;   // DC SUPPLY ON PSCB 2
   "Carrier_07_SpareInput(4_5)" AT %I716.5 : Bool;   // SPARE INPUT
   "Carrier_07_SpareInput(4_6)" AT %I716.6 : Bool;   // SPARE INPUT
   "Carrier_07_SpareInput(4_7)" AT %I716.7 : Bool;   // SPARE INPUT
   "Carrier_07_PB1_ProdHoldLH" AT %I717.0 : Bool;   // PB 1 PRODUCTION HOLD LH
   "Carrier_07_PB2_ResetLH" AT %I717.1 : Bool;   // PB 2 RESET LH
   "Carrier_07_PB3_ProdHoldRH" AT %I717.2 : Bool;   // PB 3 PRODUCTION HOLD RH
   "Carrier_07_PB4_ResetRH" AT %I717.3 : Bool;   // PB 4 RESET RH
   "Carrier_07_SpareInput(4_14)" AT %I717.4 : Bool;   // SPARE INPUT
   "Carrier_07_SpareInput(4_15)" AT %I717.5 : Bool;   // SPARE INPUT
   "Carrier_07_SpareInput(4_16)" AT %I717.6 : Bool;   // SPARE INPUT
   "Carrier_07_SpareInput(4_17)" AT %I717.7 : Bool;   // SPARE INPUT
   "Carrier_07_Slot5_Output" AT %IW718 : Word;   // SLOT 5 OUTPUT WORD
   "Carrier_07_IRD400_HMI_24VDC_ENABLE" AT %I718.0 : Bool;   // IRD 400 PANEL HMI 24V DC POWER
   "Carrier_07_FaultLight_LH" AT %I718.1 : Bool;   // FAULT LIGHT LH
   "Carrier_07_RunLight_LH" AT %I718.2 : Bool;   // RUN LIGHT LH
   "Carrier_07_FaultLight_RH" AT %I718.3 : Bool;   // FAULT LIGHT RH
   "Carrier_07_RunLight_RH" AT %I718.4 : Bool;   // RUN LIGHT RH
   "Carrier_07_SpareOutput(5_5)" AT %I718.5 : Bool;   // SPARE OUTPUT
   "Carrier_07_SpareOutput(5_6)" AT %I718.6 : Bool;   // SPARE OUTPUT
   "Carrier_07_SpareOutput(5_7)" AT %I718.7 : Bool;   // SPARE OUTPUT
   "Carrier_07_ActualSpeed" AT %IW720 : Word;   // ACTUAL SPEED
   "Carrier_07_CarrierDriveAlarm" AT %IW722 : Word;   // CARRIER DRIVE ALARM
   "Carrier_07_CarrierDriveWarning" AT %IW724 : Word;   // CARRIER DRIVE WARNING
   "Carrier_08_Status" AT %IW750 : Word;   // CARRIER STATUS WORD
   "Carrier_08_Status.0" AT %I750.0 : Bool;   // HEARTBEAT
   "Carrier_08_Status.1" AT %I750.1 : Bool;   // MANUAL
   "Carrier_08_Status.2" AT %I750.2 : Bool;   // IN_AUTO
   "Carrier_08_Status.3" AT %I750.3 : Bool;   // POSITIONING_COMPLETE
   "Carrier_08_Status.4" AT %I750.4 : Bool;   // PRODUCTION HOLD
   "Carrier_08_Status.5" AT %I750.5 : Bool;   // CARRIER MOVING FORWARD
   "Carrier_08_Status.6" AT %I750.6 : Bool;   // CARRIER MOVING REVERSE
   "Carrier_08_Status.7" AT %I750.7 : Bool;   // CARRIER FAULT
   "Carrier_08_Status.8" AT %I751.0 : Bool;   // CRASH DETECT TRIPPED
   "Carrier_08_Status.9" AT %I751.1 : Bool;
   "Carrier_08_Status.10" AT %I751.2 : Bool;
   "Carrier_08_Status.11" AT %I751.3 : Bool;
   "Carrier_08_Status.12" AT %I751.4 : Bool;
   "Carrier_08_Status.13" AT %I751.5 : Bool;
   "Carrier_08_Status.14" AT %I751.6 : Bool;
   "Carrier_08_Status.15" AT %I751.7 : Bool;
   "Carrier_08_SDCFaultCode" AT %IW752 : Word;   // SDC FAULT CODE
   "Carrier_08_CarrierPosition" AT %ID754 : DWord;   // CARRIER POSITION
   "Carrier_08_CarrierNumber" AT %IW758 : Word;   // CARRIER NUMBER
   "Carrier_08_G120DControlWord" AT %IW760 : Word;   // G120D_STW1_CONTROL
   "Carrier_08_G120DControlWord.0" AT %I760.0 : Bool;   // Bit_00_ON
   "Carrier_08_G120DControlWord.1" AT %I760.1 : Bool;   // Bit_01_AUS2_INH
   "Carrier_08_G120DControlWord.2" AT %I760.2 : Bool;   // Bit_02_AUS3_STOP
   "Carrier_08_G120DControlWord.3" AT %I760.3 : Bool;   // Bit_03_EN
   "Carrier_08_G120DControlWord.4" AT %I760.4 : Bool;   // Bit_04_EN_RAMP
   "Carrier_08_G120DControlWord.5" AT %I760.5 : Bool;   // Bit_05_START_RAMP
   "Carrier_08_G120DControlWord.6" AT %I760.6 : Bool;   // Bit_06_SETPOINT
   "Carrier_08_G120DControlWord.7" AT %I760.7 : Bool;   // Bit_07_RESET
   "Carrier_08_G120DControlWord.8" AT %I761.0 : Bool;   // Bit_08_JOG_R
   "Carrier_08_G120DControlWord.9" AT %I761.1 : Bool;   // Bit_09_JOG_L
   "Carrier_08_G120DControlWord.10" AT %I761.2 : Bool;   // Bit_10_CONTR_PLC
   "Carrier_08_G120DControlWord.11" AT %I761.3 : Bool;   // Bit_11_REVERSE
   "Carrier_08_G120DControlWord.12" AT %I761.4 : Bool;   // Bit_12_BRAKE_RELEASE
   "Carrier_08_G120DControlWord.13" AT %I761.5 : Bool;   // Bit_13_DDS
   "Carrier_08_G120DControlWord.14" AT %I761.6 : Bool;   // Bit_14_DO0
   "Carrier_08_G120DControlWord.15" AT %I761.7 : Bool;   // Bit_15_DO1
   "Carrier_08_G120DStatusWord" AT %IW762 : Word;   // G120D_ZSW1_STATUS
   "Carrier_08_G120DStatusWord.0" AT %I762.0 : Bool;   // Bit_00_READY_RUN
   "Carrier_08_G120DStatusWord.1" AT %I762.1 : Bool;   // Bit_01_READY_ON
   "Carrier_08_G120DStatusWord.2" AT %I762.2 : Bool;   // Bit_02_ENABLE